(* Logix 5000 project; controller PLC_MCC1300_75F1 vendor 1 type 14 code 166 rev 32.11; software revision 32.04; part 8 of 83 *)

        .rgxMan.4   // Run both
        .rgxMan.5   // Reverse both
        .dErrorCode2   // Error code M2
        .xSensorPresence1   // M403.P115B1.Synchro photocell / start count {x|x|x|x|O}
        .xSensorPresence2   // M403.P115B2.Synchro photocell / start count {x|x|x|x|O}
   M311_HMW : MAC_Conveyor_HMW;
        .dParam_1_cmm   // Positioning offset 1 [mm] {mm/100|mm|-50|+50|M}
        .dParam_2_cmm   // Positioning offset 2 [mm] {mm/100|mm|-50|+50|M}
        .rgxMan.0   // Run M1
        .rgxMan.1   // Reverse M1
        .rgxMan.2   // Run M2
        .rgxMan.3   // Reverse M2
        .rgxMan.4   // Run both
        .rgxMan.5   // Reverse both
   M311_M1_DR : AXIS_CIP_DRIVE; {access Read Only}
   M311_M1_DR_IN_MAJ : MOTION_INSTRUCTION := (FLAGS := 570425344, DN := 1); {access None}
   M311_M1_DR_IN_MAM : MOTION_INSTRUCTION := (FLAGS := 704643072, DN := 1, PC := 1); {access None}
   M311_M1_DR_IN_MAR : MOTION_INSTRUCTION := (FLAGS := 167772160, PC := 1); {access None}
   M311_M1_DR_IN_MAS : MOTION_INSTRUCTION := (FLAGS := -1442840576, EN := 1, DN := 1, PC := 1); {access None}
   M311_M1_DR_IN_MCD : MOTION_INSTRUCTION := (FLAGS := 570425344, DN := 1); {access None}
   M311_M1_DR_IN_MRP : MOTION_INSTRUCTION := (FLAGS := 536870912, DN := 1, STATUS := 2, STATE := 3); {access None}
   M311_M1_DR_MAFR : MOTION_INSTRUCTION := (FLAGS := 301989888, ER := 1, ERR := 11); {access None}
   M311_M1_DR_MDR : MOTION_INSTRUCTION := (FLAGS := -1845493760, EN := 1, ER := 1, ERR := 11); {access None}
   M311_M1_DR_MSF : MOTION_INSTRUCTION := (FLAGS := 570425344, DN := 1, STATUS := 2, STATE := 1); {access None}
   M311_M1_DR_MSO : MOTION_INSTRUCTION := (FLAGS := -1610612736, EN := 1, DN := 1, STATE := 1); {access None}
   M311_M1_DR_OUT_MAJ : MOTION_INSTRUCTION := (FLAGS := 570425344, DN := 1); {access None}
   M311_M1_DR_OUT_MAM : MOTION_INSTRUCTION := (FLAGS := 704643072, DN := 1, PC := 1); {access None}
   M311_M1_DR_OUT_MAR : MOTION_INSTRUCTION := (FLAGS := 671088640, DN := 1, PC := 1, STATE := 1); {access None}
   M311_M1_DR_OUT_MAS : MOTION_INSTRUCTION := (FLAGS := -1442840576, EN := 1, DN := 1, PC := 1); {access None}
   M311_M1_DR_OUT_MCD : MOTION_INSTRUCTION := (FLAGS := 570425344, DN := 1); {access None}
   M311_M1_DR_OUT_MRP : MOTION_INSTRUCTION := (FLAGS := 536870912, DN := 1, STATUS := 2, STATE := 3); {access None}
   M311_SpaceConv_Utilities : SpaceConv_Utilities := (CONST_dSyncMode := 1, CONST_dSyncroPhWindow_cmm := 450000, CONST_dConveyorLength_cmm := 800000, CONST_dConveyorWidth_cmm := 400000, CONST_dPresetFeedbackTime_ms := 500, CONST_rAcceleration_ms2 := 1.2, CONST_rDeceleration_ms2 := 1.2, CONF_MD1_dScan_ms := 20, CONF_MD2_MD3_dPrstPos_cmm := -390000, CONF_MD4_MD6_dLength_cmm := 365800, CONF_MD7_dOffset_cmm := 50000, ST_dStopLoadForseen_cmm := 620000, ST_dRealSpeed_mm_min := 90000, ST_rStepAdvancementH := 3000.0, ST_rStepAdvancementT := 3000.0, O_xPlateSynchronized := 1, O_dCountFeedbackTime_ms := 500, O_dPresetLoadUnload_cmm := -126300);
   M311_SpaceConvUtilities : SpaceConv_Utilities; {access Read Only}
   M311_TON_Synchro_timeout : TIMER; {access Read Only}
   M311_xOS_SentToCullet : BOOL; {access Read Only}
   M311_xPlateCullet : BOOL; {access Read Only}
   M311_xSendCulletReqActive : BOOL; {access Read Only}
   M311_xSensorTimeout : BOOL; {access Read Only}
   M311A : MAC_Rotator := (ST_xCleaningConditionOK := 1, ST_xConditionOKStopCycle := 1, ST_xEnableControlError := 1, INPUT_rRotatorPosition_cdeg := 26999.898, INPUT_xConditionToDescent := 1, INPUT_xLowPosition := 1, INPUT_xLocalSafetySwitchRotation := 1, INPUT_xProtectionMotorLifting := 1, INPUT_xProtectionMotorRotation := 1, tmON_DelayFrameUP.PRE := 100, tmON_DelayRotatorInRun.PRE := 300, tmOF_DriveEnable.PRE := 20000, tmOF_DriveEnable.ACC := 20000, tmON_FeedbackTimeOutLifting.PRE := 1000, tmON_FeedbackTimeOutRotation.PRE := 1000, tmON_FramePosError.PRE := 2500, tmON_RotatePosError.PRE := 10000, tmON_RotatePosError.ACC := 2040, tmON_RotatePosError.EN := 1, tmON_RotatePosError.TT := 1, tmON_PresetEncoder.PRE := 3000, tmON_DelayBrakeON.PRE := 200); {access None}
        .OUTPUT_xDescent   // P253KA4.Descent frame
        .PH_x.0   // Rise frame
        .PH_x.12   // Counterclockwise rotation
        .PH_x.4   // Descent frame
        .PH_x.8   // Clockwise totation
        .OUTPUT_xRise   // P253KA3.Lifting frame
        .INPUT_xLowPosition   // P56KA2.Frame to low position
        .INPUT_xFeedbackLifting   // P56KM1/2.Feedback lifting chassis
        .INPUT_xHighPosition   // P56KA1.Frame to high position
        .INPUT_xProtectionMotorLifting   // P56QM1.Protection lifting frame
   M311A_ALM : MAC_Rotator_ALM;
        .rgxStoppingFault_M[0].0   // Z401.M311A.Protection motor rotation
        .rgxStoppingFault_M[0].1   // Z401.M311A.Drive Error
        .rgxStoppingFault_M[0].11   // Z401.M311A.Frame lifting position error
        .rgxStoppingFault_M[0].2   // Z401.M311A.Drive feedback error
        .rgxStoppingFault_M[0].20   // Z401.M311A.Drive not ready
        .rgxStoppingFault_M[0].3   // Z401.M311A.Rotation position error
        .rgxStoppingFault_M[0].8   // Z401.M311A.Protection lifting frame
        .rgxStoppingFault_M[0].9   // Z401.M311A.Feedback lifting chassis
   M311A_Data : UDT_Convoy_SL;
   M311A_HMR : MAC_Rotator_HMR := (xLowPosition := 1, dState := 1, dActualAngle_cdeg := 27000);
        .rgxMan.0   // Rise
        .rgxMan.1   // Descent
        .rgxMan.10   // Clockwise rotation jog
        .rgxMan.11   // Counter Clockwise rotation jog
        .rgxMan.14   // Enable brake release
        .rgxMan.15   // Disable brake release
        .rgxMan.8   // Clockwise rotation
        .rgxMan.9   // Counter Clockwise rotation
   M311A_HMW : MAC_Rotator_HMW := (xPresetEnc := 1, dLowSpeed_deg_s := 40, dLowRamp_deg_s2 := 50, dHighSpeed_deg_s := 50, dHighRamp_deg_s2 := 60, dJogSpeed_deg_s := 12);
        .rgxMan.0   // Rise
        .rgxMan.1   // Descent
        .rgxMan.10   // Clockwise rotation jog
        .rgxMan.11   // Counterclockwise rotation jog
        .rgxMan.14   // Enable brake release
        .rgxMan.15   // Disable brake release
        .rgxMan.8   // Clockwise rotation
        .rgxMan.9   // Counterclockwise rotation
   M311A_M1_DR : AXIS_CIP_DRIVE; {access Read Only}
   M311A_M1_DR_IN_MAJ : MOTION_INSTRUCTION := (FLAGS := 570425344, DN := 1); {access None}
   M311A_M1_DR_IN_MAM : MOTION_INSTRUCTION := (FLAGS := 704643072, DN := 1, PC := 1); {access None}
   M311A_M1_DR_IN_MAS : MOTION_INSTRUCTION := (FLAGS := -1442840576, EN := 1, DN := 1, PC := 1); {access None}
   M311A_M1_DR_MAFR : MOTION_INSTRUCTION := (FLAGS := 301989888, ER := 1, ERR := 11); {access None}
   M311A_M1_DR_MAH : MOTION_INSTRUCTION := (FLAGS := 671088640, DN := 1, PC := 1, STATE := 17); {access None}
   M311A_M1_DR_MSF : MOTION_INSTRUCTION := (FLAGS := -1610612736, EN := 1, DN := 1, STATUS := 2, STATE := 1); {access None}
   M311A_M1_DR_MSO : MOTION_INSTRUCTION := (FLAGS := 536870912, DN := 1, STATE := 1); {access None}
   M311A_M1_DR_OUT_MAJ : MOTION_INSTRUCTION := (FLAGS := 570425344, DN := 1); {access None}
   M311A_M1_DR_OUT_MAM : MOTION_INSTRUCTION := (FLAGS := 704643072, DN := 1, PC := 1); {access None}
   M311A_M1_DR_OUT_MAS : MOTION_INSTRUCTION := (FLAGS := -1442840576, EN := 1, DN := 1, PC := 1); {access None}
   M311A_MAM_IP_TOFF : TIMER; {access Read Only}
   M311A_rLastPosition : REAL; {access Read Only}
   M311A_TmON1 : TIMER; {access Read Only}
   M311M312_OffsetBaricentre_cmm : DINT; {access Read Only}
   M312 : MAC_Conveyor_Single := (ST_xCleaningConditionOK := 1, ST_xPlatePresence := 1, ST_xConditionOKStopCycle := 1, ST_xOutputEnable := 1, ST_xIdPlatePresence := 1, ST_xWaitStopNextMachine := 1, ST_xEnableControlError := 1, ST_xPlateSynchronized := 1, ST_xSafetyMovement := 1, OSR_xSynchroPhotocellTail := 1, INPUT_xSquaringPhotocell_4 := 1, INPUT_xLowPositionSquaring_1 := 1, INPUT_xHighPositionPopup_1 := 1, INPUT_xHighPositionPopup_2 := 1, INPUT_xDriveReady_M1 := 1, INPUT_xLocalSafetySwitch_M1 := 1, INPUT_xMotorThermalProbe_M1 := 1, INPUT_xProtectionMotor_M1 := 1, INPUT_xDriveReady_M2 := 1, INPUT_xLocalSafetySwitch_M2 := 1, INPUT_xMotorThermalProbe_M2 := 1, INPUT_xProtectionMotor_M2 := 1, INPUT_xDriveFeedback_M3 := 1, INPUT_xDriveReady_M3 := 1, INPUT_xLocalSafetySwitch_M3 := 1, INPUT_xMotorThermalProbe_M3 := 1, INPUT_xProtectionMotor_M3 := 1, INPUT_xDriveReady_M4 := 1, INPUT_xLocalSafetySwitch_M4 := 1, INPUT_xMotorThermalProbe_M4 := 1, INPUT_xProtectionMotor_M4 := 1, INPUT_xProtectionLiftingFrame_1 := 1, INPUT_xProtectionLiftingFrame_2 := 1, INPUT_xFeedbackVentilation_1 := 1, INPUT_xFeedbackVentilation_2 := 1, OUTPUT_xDriveEnable_M1 := 1, OUTPUT_xDriveEnable_M2 := 1, OUTPUT_xDriveEnable_M3 := 1, OUTPUT_xDriveEnable_M4 := 1, OUTPUT_xFunCommand_1 := 1, OUTPUT_xFunCommand_2 := 1, AUX_dPresetStopLoad_cmm := 372333, AUX_dPresetStopUnload_cmm := 441667, AUX_dAccSpace_cmm := 41667, AUX_dDecSpace_cmm := 41667, AUX_dReqSpeed_mm_min := 60000, AUX_dAbsPosTarget_M3_cmm := 195500, AUX_dAbsPosTarget_M4_cmm := 195500, AUX_dQtaLites := 1, tmON_FeedbackTimeOut_M1.PRE := 2000, tmOF_DriveEnable_M1.PRE := 30000, tmOF_DriveEnable_M1.ACC := 540, tmOF_DriveEnable_M1.TT := 1, tmOF_DriveEnable_M1.DN := 1, tmOF_PowerSaving_M1.EN := 1, tmOF_PowerSaving_M1.DN := 1, tmON_FeedbackTimeOut_M2.PRE := 2000, tmOF_DriveEnable_M2.PRE := 30000, tmOF_DriveEnable_M2.ACC := 540, tmOF_DriveEnable_M2.TT := 1,
        tmOF_DriveEnable_M2.DN := 1, tmON_FeedbackTimeOut_M3.PRE := 2000, tmOF_DriveEnable_M3.PRE := 30000, tmOF_DriveEnable_M3.ACC := 540, tmOF_DriveEnable_M3.TT := 1, tmOF_DriveEnable_M3.DN := 1, tmON_FeedbackTimeOut_M4.PRE := 2000, tmOF_DriveEnable_M4.PRE := 30000, tmOF_DriveEnable_M4.ACC := 540, tmOF_DriveEnable_M4.TT := 1, tmOF_DriveEnable_M4.DN := 1, tmON_AuxFunction1.PRE := 5000, tmON_AuxFunction1.EN := 1, tmON_AuxFunction1.DN := 1, tmON_AuxFunction2.PRE := 2200, tmON_AuxFunction3.PRE := 2200, tmON_AuxFunction4.PRE := 15000, tmON_AuxFunction5.PRE := 3000, tmON_AuxFunction6.PRE := 15000, tmON_AuxFunction7.PRE := 3600000, tmON_AuxFunction8.PRE := 40000, tmON_AuxFunction9.PRE := 20000, TmON[0].PRE := 3000, TmON[1].PRE := 1000, TmON[1].ACC := 1019, TmON[2].PRE := 5000, TmON[6].PRE := 5000, TmON[6].EN := 1, TmON[6].DN := 1, TmON[11].PRE := 2000, TmON[12].PRE := 2000, TmON[13].PRE := 2000, TmON[14].PRE := 2000, tmOF_MCD_M1.ACC := 20, tmOF_MCD_M2.ACC := 20, tmOF_MCD_M3.ACC := 20, tmOF_MCD_M4.ACC := 20); {access None}
        .INPUT_xSquaringPhotocell_1   // P406B1.Squaring frontal photocell - Right
        .INPUT_xMotorThermalProbe_M2   // M2.P404BT2.Motor thermal probe
        .INPUT_xLowPositionPopup_1   // P63KA2.M5.Low position popup
        .INPUT_xLowPositionSquaring_1   // P405SQ2.Low position squaring
        .INPUT_xMotorThermalProbe_M1   // M1.P404BT1.Motor thermal probe
        .INPUT_xHighPositionPopup_1   // P63KA1.M5.High position popup
        .INPUT_xSquaringPhotocell_2   // P406B2.Squaring frontal photocell - Left
        .INPUT_xHighPositionPopup_2   // P64KA1.M6.High position popup
        .PH_x.0   // Load (from M311)
        .PH_x.10   // Load (from M409)
        .PH_x.11   // End load (from M409)
        .PH_x.12   // Unload (to M311)
        .PH_x.13   // End unload (to M311)
        .PH_x.15   // End unload (to M409)
        .PH_x.16   // Rise popup
        .PH_x.19   // End rise popup
        .PH_x.20   // Descent popup
        .PH_x.23   // End descent popup
        .PH_x.24   // Reset counter position
        .PH_x.26   // Lateral positioning (M3-M4)
        .PH_x.27   // End lateral positioning (M3-M4)
        .PH_x.28   // Lateral squaring
        .PH_x.29   // End lateral squaring
        .PH_x.30   // Lateral traction recovery (M3-M4)
        .PH_x.31   // End lateral traction recovery (M3-M4)
        .PH_x.4   // Frontal squaring (run fwd + rise squaring)
        .PH_x.5   // End frontal sqauring
        .PH_x.7   // End load (from M311)
        .PH_x.8   // Unload (to M409)
        .INPUT_xMotorThermalProbe_M3   // M3.P405BT3.Motor thermal probe
        .INPUT_xLowPositionPopup_2   // P64KA2.M6.Low position popup
        .INPUT_xSquaringPhotocell_3   // P405B1.Squaring lateral photocell - Right
        .INPUT_xHighPositionSquaring_1   // P405SQ1.High position squaring
        .INPUT_xSquaringPhotocell_4   // P405B2.Squaring lateral photocell - Left
        .INPUT_xHighPositionSquaring_2   // P405SQ11.High position squaring
        .ST_xAux1   // Ready to unload on backward conveyor
        .INPUT_xLowPositionSquaring_2   // P405SQ12.Low position squaring
   M312_ALM : MAC_Conveyor_ALM;
        .rgdFaultCode_M[0]   // Drive fault code M1
        .rgdFaultCode_M[1]   // Drive fault code M2
        .rgxStoppingFault[0].0   // Z401.M312-M1.Positioning error
        .rgxStoppingFault[0].1   // Z401.M312-M1.Plate not synchronized
        .rgxStoppingFault[0].10   // Z401.M312-M2.Error position frontal squaring
        .rgxStoppingFault[0].11   // Z401.M312-M2.Timeout frontal squaring
        .rgxStoppingFault[0].12   // Z401.M312-M2.Lugs position sensors fault
        .rgxStoppingFault[0].13   // Z401.M312.Timeout movement popup 1
        .rgxStoppingFault[0].14   // Z401.M312.Timeout movement popup 1
        .rgxStoppingFault[0].16   // Z401.M312-M3.Positioning error
        .rgxStoppingFault[0].18   // Z401.M312-M3.Error position popup
        .rgxStoppingFault[0].19   // Z401.M312-M3.Error position lateral squaring
        .rgxStoppingFault[0].2   // Z401.M312-M1.Error position frontal squaring
        .rgxStoppingFault[0].20   // Z401.M312-M3.Timeout lateral squaring
        .rgxStoppingFault[0].21   // Z401.M312.Protection lifting popup 1
        .rgxStoppingFault[0].22   // Z401.M312.Protection lifting popup 2
        .rgxWarning[0].10   // Z401.M312_M2.Plate not synchronized
        .rgxStoppingFault[0].3   // Z401.M312-M1.Timeout frontal squaring
        .rgxStoppingFault[0].4   // Z401.M312-M1.Lugs position sensors fault
        .rgxStoppingFault[0].5   // Z401.M312.Popup 1 position error
        .rgxStoppingFault[0].6   // Z401.M312.Popup 2 position error
        .rgxStoppingFault[0].8   // Z401.M312-M2.Positioning error
        .rgxStoppingFault[0].9   // Z401.M312-M2.Plate not synchronized
        .rgxStoppingFault_M[0].0   // Z401.M312-M1.Protection motor rotation
        .rgxStoppingFault_M[0].1   // Z401.M312-M1.Drive error
        .rgxStoppingFault_M[0].10   // Z401.M312-M2.Drive feedback error
        .rgxStoppingFault_M[0].11   // Z401.M312-M2.Local safety switch
        .rgxStoppingFault_M[0].12   // Z401.M312-M2.Motor thermal probe
        .rgxStoppingFault_M[0].13   // Z401.M312-M2.Braking resistor anomaly
        .rgxStoppingFault_M[0].14   // Z401.M312-M2.Drive not ready
        .rgxStoppingFault_M[0].16   // Z401.M312-M3.Protection motor rotation
        .rgxStoppingFault_M[0].17   // Z401.M312-M3.Drive error
        .rgxStoppingFault_M[0].18   // Z401.M312-M3.Drive feedback error
        .rgxStoppingFault_M[0].19   // Z401.M312-M3.Local safety switch
        .rgxStoppingFault_M[0].2   // Z401.M312-M1.Drive feedback error
        .rgxStoppingFault_M[0].20   // Z401.M312-M3.Motor thermal probe
        .rgxStoppingFault_M[0].21   // Z401.M312-M3.Drive not ready
        .rgxStoppingFault_M[0].3   // Z401.M312-M1.Local safety switch
        .rgxStoppingFault_M[0].4   // Z401.M312-M1.Motor thermal probe
        .rgxStoppingFault_M[0].5   // Z401.M312-M1.Braking resistor anomaly
        .rgxStoppingFault_M[0].6   // Z401.M312-M1.Drive not ready
        .rgxStoppingFault_M[0].8   // Z401.M312-M2.Protection motor rotation
        .rgxStoppingFault_M[0].9   // Z401.M312-M2.Drive error
        .rgxWarning[0].0   // Z401.M312_M1.Plate not synchronized
        .rgxWarning[0].1   // Z401.M312_M1.Positioning error
        .rgxWarning[0].11   // Z401.M312_M2.Positioning error
        .rgxWarning[0].21   // Z401.M312_M3.Lateal positioning error
        .rgxWarning[0].25   // Z401.M312.Timeout frontal squaring
        .rgxWarning[0].26   // Z401.M312.Timeout lateral squaring
   M312_AlmTimer1 : TIMER; {access Read Only}
   M312_AlmTimer2 : TIMER; {access Read Only}
   M312_Data : UDT_Convoy_SL;
        .rgtCap[0].rgxRequest.0   // Frontal squaring request
        .rgtCap[0].rgxRequest.1   // Lateral squaring request
        .rgtCap[0].rgxRequest.2   // Y adjust position request
        .rgtCap[0].rgxRequest.3   // Y measure request
        .rgtCap[0].rgxDone.0   // Frontal squaring done
        .rgtCap[0].rgxDone.1   // Lateral squaring done
        .rgtCap[0].rgxDone.2   // Y adjust position done
        .rgtCap[0].rgxDone.3   // Y measure done
   M312_dSlowingSquaringQuote : DINT; {access Read Only}
   M312_dTractionRecovery_M3 : DINT; {access Read Only}
   M312_dTractionRecovery_M4 : DINT; {access Read Only}
   M312_HMR : MAC_Conveyor_HMR := (xSensorPresence4 := 1, xHighPositionPopup1 := 1, xHighPositionPopup2 := 1, xLowPositionSquaring1 := 1, xLowPositionSquaring2 := 1, xIdPlatePresence := 1, dState1 := 1, dState2 := 1, dState3 := 1, dState4 := 1, dStateSensor1 := 1, dStateSensor2 := 1, dStateSensor3 := 1, dStateSensor4 := 1, dStateSensor5 := 1, dStateSensor6 := 1);
        .xSensorPresence5   // P115/3.Start count photocell {x|x|x|x|O}
        .xHighPositionPopup2   // P64KA1.M6.High position popup {x|x|x|x|O}
        .dErrorCode1   // Error code M1
        .xHighPositionPopup1   // P63KA1.M5.High position popup {x|x|x|x|O}
        .rgxMan.0   // Run M1
        .rgxMan.1   // Reverse M1
        .rgxMan.10   // Rise popup 1
        .rgxMan.11   // Descent popup 1
        .rgxMan.12   // Rise popup 2
        .rgxMan.13   // Descent popup 2
        .rgxMan.14   // Rise all popups
        .rgxMan.15   // Descent all popups
        .rgxMan.16   // Rise frontal squaring 1
        .rgxMan.17   // Descent frontal squaring 1
        .rgxMan.18   // Rise frontal squaring 2
        .rgxMan.19   // Descent frontal squaring 2
        .rgxMan.2   // Run M2
        .rgxMan.20   // Rise all frontal squaring
        .rgxMan.21   // Descent all frontal squaring
        .rgxMan.3   // Reverse M2
        .rgxMan.4   // Run M3
        .rgxMan.5   // Reverse M3
        .rgxMan.6   // Run M4
        .rgxMan.7   // Reverse M4
        .dState3   // State M3 (1=No anomaly; 3=Run; 4=Reverse; 7=Anomaly)
        .xHighPositionSquaring1   // P405SQ1.High position frontal squaring M1 {x|x|x|x|O}
        .dErrorCode2   // Error code M2
        .xSensorPresence6   // P115/4.Start count photocell {x|x|x|x|O}
        .xSensorPresence4   // P404B1.SlowDown photocell frontal squaring left {x|x|x|x|O}
        .xLowPositionPopup1   // P63KA2.M5.Low position popup {x|x|x|x|O}
        .xHighPositionSquaring2   // P405SQ11.High position frontal squaring M2 {x|x|x|x|O}
        .dState2   // State M2 (1=No anomaly; 3=Run; 4=Reverse; 7=Anomaly)
        .dErrorCode4   // Error code M4
        .xSensorPresence3   // P404B1.SlowDown photocell frontal squaring right {x|x|x|x|O}
        .dState1   // State M1 (1=No anomaly; 3=Run; 4=Reverse; 7=Anomaly)
        .dState4   // State M4 (1=No anomaly; 3=Run; 4=Reverse; 7=Anomaly)
        .xLowPositionSquaring2   // P405SQ12.Low position frontal squaring M2 {x|x|x|x|O}
        .xLowPositionSquaring1   // P405SQ2.Low position frontal squaring M1 {x|x|x|x|O}
        .xLowPositionPopup2   // P64KA2.M6.Low position popup {x|x|x|x|O}
        .xSensorPresence1   // P405B1.SlowDown photocell lateral squaring right {x|x|x|x|O}
        .dErrorCode3   // Error code M3
        .xSensorPresence2   // P405B2.SlowDown photocell lateral squaring left {x|x|x|x|O}
   M312_HMW : MAC_Conveyor_HMW := (dParam_3_cmm := 4000, dParam_5_ms := 3000, dParam_6_ms := 4000, dParam_7_ms := 2200, dParam_8_ms := 5000);
        .dParam_4_cmm   // Lateral squaring space {mm/100|mm|0|500|M}
        .dParam_1_cmm   // Positioning offset 1 {mm/100|mm|-50|+50|M}
        .dParam_3_cmm   // Frontal squaring space {mm/100|mm|0|500|M}
        .dParam_6_ms   // Squaring frontal time 2 {ms|s|0|5|M}
        .dParam_2_cmm   // Positioning offset 2 {mm/100|mm|-50|+50|M}
        .dParam_8_ms   // Squaring lateral time 2 {ms|s|0|5|M}
        .rgxMan.0   // Run M1
        .rgxMan.1   // Reverse M1
        .rgxMan.10   // Rise popup 2
        .rgxMan.11   // Descent popup 2
        .rgxMan.12   // Rise all popups
        .rgxMan.13   // Descent all popups
        .rgxMan.14   // Run both (M1-2)
        .rgxMan.15   // Reverse both (M1-2)
        .rgxMan.16   // Rise frontal squaring 1
        .rgxMan.17   // Descent frontal squaring 1
        .rgxMan.18   // Rise frontal squaring 2
        .rgxMan.19   // Descent frontal squaring 2
        .rgxMan.2   // Run M2
        .rgxMan.20   // Rise all frontal squaring
        .rgxMan.21   // Descent all frontal squaring
        .rgxMan.3   // Reverse M2
        .rgxMan.4   // Run M3
        .rgxMan.5   // Reverse M3
        .rgxMan.6   // Run M4
        .rgxMan.7   // Reverse M4
        .rgxMan.8   // Rise popup 1
        .rgxMan.9   // Descent popup 1
        .dParam_7_ms   // Squaring lateral time 1 {ms|s|0|5|M}
        .dParam_5_ms   // Squaring frontal time 1 {ms|s|0|5|M}
   M312_M1_DR_IN_MAJ : MOTION_INSTRUCTION := (FLAGS := 570425344, DN := 1); {access None}
   M312_M1_DR_IN_MAM : MOTION_INSTRUCTION := (FLAGS := 33554432); {access None}
   M312_M1_DR_IN_MAR : MOTION_INSTRUCTION := (FLAGS := 33554432); {access None}
   M312_M1_DR_IN_MAS : MOTION_INSTRUCTION := (FLAGS := -1442840576, EN := 1, DN := 1, PC := 1); {access None}
   M312_M1_DR_IN_MCD : MOTION_INSTRUCTION := (FLAGS := 570425344, DN := 1); {access None}
   M312_M1_DR_IN_MRP : MOTION_INSTRUCTION := (FLAGS := 33554432); {access None}
   M312_M1_DR_MAFR : MOTION_INSTRUCTION := (FLAGS := 301989888, ER := 1, ERR := 11); {access None}
   M312_M1_DR_MDR : MOTION_INSTRUCTION := (FLAGS := -1845493760, EN := 1, ER := 1, ERR := 11); {access None}
   M312_M1_DR_MSF : MOTION_INSTRUCTION := (FLAGS := 570425344, DN := 1, STATUS := 2, STATE := 1); {access None}
   M312_M1_DR_MSO : MOTION_INSTRUCTION := (FLAGS := -1610612736, EN := 1, DN := 1, STATE := 1); {access None}
   M312_M1_DR_OUT_MAJ : MOTION_INSTRUCTION := (FLAGS := 570425344, DN := 1); {access None}
   M312_M1_DR_OUT_MAM : MOTION_INSTRUCTION := (FLAGS := 33554432); {access None}
   M312_M1_DR_OUT_MAR : MOTION_INSTRUCTION := (FLAGS := 33554432); {access None}
   M312_M1_DR_OUT_MAS : MOTION_INSTRUCTION := (FLAGS := -1442840576, EN := 1, DN := 1, PC := 1); {access None}
   M312_M1_DR_OUT_MCD : MOTION_INSTRUCTION := (FLAGS := 570425344, DN := 1); {access None}
   M312_M1_DR_OUT_MRP : MOTION_INSTRUCTION := (FLAGS := 33554432); {access None}
   M312_M1_DR_R1 : AXIS_CIP_DRIVE; {access Read Only}
   M312_M2_AUX_ReqSpeed_mm_min : DINT; {access Read Only}
   M312_M2_ChangeSpeed : BOOL; {access Read Only}
   M312_M2_DR_IN_MAJ : MOTION_INSTRUCTION := (FLAGS := 570425344, DN := 1); {access None}
   M312_M2_DR_IN_MAM : MOTION_INSTRUCTION := (FLAGS := 33554432); {access None}
   M312_M2_DR_IN_MAR : MOTION_INSTRUCTION := (FLAGS := 33554432); {access None}
   M312_M2_DR_IN_MAS : MOTION_INSTRUCTION := (FLAGS := 704643072, DN := 1, PC := 1); {access None}
   M312_M2_DR_IN_MCD : MOTION_INSTRUCTION := (FLAGS := 301989888, ER := 1, ERR := 23); {access None}
   M312_M2_DR_IN_MRP : MOTION_INSTRUCTION := (FLAGS := 536870912, DN := 1, STATUS := 2, STATE := 3); {access None}
   M312_M2_DR_MAFR : MOTION_INSTRUCTION := (FLAGS := 301989888, ER := 1, ERR := 11); {access None}
   M312_M2_DR_MDR : MOTION_INSTRUCTION := (FLAGS := -1845493760, EN := 1, ER := 1, ERR := 11); {access None}
   M312_M2_DR_MSF : MOTION_INSTRUCTION := (FLAGS := 570425344, DN := 1, STATUS := 2, STATE := 1); {access None}
   M312_M2_DR_MSO : MOTION_INSTRUCTION := (FLAGS := -1610612736, EN := 1, DN := 1, STATE := 1); {access None}
   M312_M2_DR_OUT_MAJ : MOTION_INSTRUCTION := (FLAGS := 570425344, DN := 1); {access None}
   M312_M2_DR_OUT_MAM : MOTION_INSTRUCTION := (FLAGS := 33554432); {access None}
   M312_M2_DR_OUT_MAR : MOTION_INSTRUCTION := (FLAGS := 33554432); {access None}
   M312_M2_DR_OUT_MAS : MOTION_INSTRUCTION := (FLAGS := 704643072, DN := 1, PC := 1); {access None}
   M312_M2_DR_OUT_MCD : MOTION_INSTRUCTION := (FLAGS := 301989888, ER := 1, ERR := 23); {access None}
   M312_M2_DR_OUT_MRP : MOTION_INSTRUCTION := (FLAGS := 536870912, DN := 1, STATUS := 2, STATE := 3); {access None}
   M312_M2_DR_R2 : AXIS_CIP_DRIVE; {access Read Only}
   M312_M2_ReqSpeed_mm_min : DINT; {access Read Only}
   M312_M3_AUX_ReqSpeed_mm_min : DINT; {access Read Only}
   M312_M3_ChangeSpeed : BOOL; {access Read Only}
   M312_M3_DR_IN_MAJ : MOTION_INSTRUCTION := (FLAGS := 570425344, DN := 1); {access None}
   M312_M3_DR_IN_MAM : MOTION_INSTRUCTION := (FLAGS := -1509949440, EN := 1, DN := 1, IP := 1); {access None}
   M312_M3_DR_IN_MAR : MOTION_INSTRUCTION := (FLAGS := 33554432); {access None}
   M312_M3_DR_IN_MAS : MOTION_INSTRUCTION := (FLAGS := 704643072, DN := 1, PC := 1); {access None}
   M312_M3_DR_IN_MCD : MOTION_INSTRUCTION := (FLAGS := 570425344, DN := 1); {access None}
   M312_M3_DR_IN_MRP : MOTION_INSTRUCTION := (FLAGS := 536870912, DN := 1, STATUS := 2, STATE := 3); {access None}
   M312_M3_DR_L : AXIS_CIP_DRIVE; {access Read Only}
   M312_M3_DR_MAFR : MOTION_INSTRUCTION := (FLAGS := 301989888, ER := 1, ERR := 11); {access None}
   M312_M3_DR_MDR : MOTION_INSTRUCTION := (FLAGS := -1845493760, EN := 1, ER := 1, ERR := 11); {access None}
   M312_M3_DR_MSF : MOTION_INSTRUCTION := (FLAGS := 570425344, DN := 1, STATUS := 2, STATE := 1); {access None}
   M312_M3_DR_MSO : MOTION_INSTRUCTION := (FLAGS := -1610612736, EN := 1, DN := 1, STATE := 1); {access None}
   M312_M3_DR_OUT_MAJ : MOTION_INSTRUCTION := (FLAGS := 570425344, DN := 1); {access None}
   M312_M3_DR_OUT_MAM : MOTION_INSTRUCTION := (FLAGS := -1509949440, EN := 1, DN := 1, IP := 1);
   M312_M3_DR_OUT_MAR : MOTION_INSTRUCTION := (FLAGS := 33554432); {access None}
   M312_M3_DR_OUT_MAS : MOTION_INSTRUCTION := (FLAGS := 704643072, DN := 1, PC := 1); {access None}
   M312_M3_DR_OUT_MCD : MOTION_INSTRUCTION := (FLAGS := 570425344, DN := 1); {access None}
   M312_M3_DR_OUT_MRP : MOTION_INSTRUCTION := (FLAGS := 536870912, DN := 1, STATUS := 2, STATE := 3); {access None}
   M312_M3_ReqSpeed_mm_min : DINT; {access Read Only}
   M312_M3_xOSR_LatSquarFtc : BOOL; {access Read Only}
   M312_SpaceConv_Utilities : SpaceConv_Utilities := (CONST_dSyncMode := 1, CONST_dSyncroPhWindow_cmm := 450000, CONST_dConveyorLength_cmm := 800000, CONST_dConveyorWidth_cmm := 400000, CONST_dPresetFeedbackTime_ms := 500, CONST_rAcceleration_ms2 := 1.2, CONST_rDeceleration_ms2 := 1.2, CONF_MD1_dScan_ms := 20, CONF_MD2_MD3_dPrstPos_cmm := -390000, CONF_MD4_MD6_dLength_cmm := 365800, CONF_MD7_dOffset_cmm := 50000, ST_dStopLoadForseen_cmm := 620000, ST_dRealSpeed_mm_min := 90000, ST_rStepAdvancementH := 3000.0, ST_rStepAdvancementT := 3000.0, O_xPlateSynchronized := 1, O_dCountFeedbackTime_ms := 500, O_dPresetLoadUnload_cmm := -126300);
   M312_TimerAlm3 : TIMER; {access Read Only}
   M312_TON_FrontSquarLeft_timeout : TIMER; {access Read Only}
   M312_TON_FrontSquarRight_timeout : TIMER; {access Read Only}
   M312_TON_LatSquarLeft_timeout : TIMER; {access Read Only}
   M312_TON_LatSquarRight_timeout : TIMER; {access Read Only}
   M312_TON_Load : TIMER; {access Read Only}
   M312_TON_Synchro_timeout : TIMER; {access Read Only}
   M312_xEnableTractionRecovering : BOOL; {access Read Only}
   M312_xFrontLeftTimeout : BOOL; {access Read Only}
   M312_xFrontRightTimeout : BOOL; {access Read Only}
   M312_xLateralTractionRecovered : BOOL; {access Read Only}
   M312_xLatLeftTimeout : BOOL; {access Read Only}
   M312_xLatRightTimeout : BOOL; {access Read Only}
   M312_xOS_PosReq : BOOL;
   M312_xPlateCullet : BOOL; {access Read Only}
   M312_xSendCulletReqActive : BOOL; {access Read Only}
   M312_xSensorTimeout : BOOL; {access Read Only}
   M315_M1_DR_R1 : AXIS_CIP_DRIVE; {access Read Only}
   M315_M2_DR_R2 : AXIS_CIP_DRIVE; {access Read Only}
   M315_M3_DR_R3 : AXIS_CIP_DRIVE; {access Read Only}
   M315_M4_DR_B1 : AXIS_CIP_DRIVE; {access Read Only}
   M315_M5_DR_B2 : AXIS_CIP_DRIVE; {access Read Only}
   M315_M6_DR_L1 : AXIS_CIP_DRIVE; {access Read Only}
   M315_M7_DR_L2 : AXIS_CIP_DRIVE; {access Read Only}
   M315_xReqStopPrevConvForPos : BOOL; {access Read Only}
   M315A : MAC_Conveyor;
        .PH_x.1   // Load Upstream
        .PH_x.0   // Load
        .PH_x.7   // End load
        .PH_x.8   // Unload
        .PH_x.15   // End unload
        .INPUT_xMotorThermalProbe_M1   // M315A.M1.Q403BT3. Motor thermal probe
        .PH_x.2   // Load Downstream
        .PH_x.5   // End load Upstream
        .PH_x.6   // End load Downstream
        .PH_x.9   // Unload Upstream
        .PH_x.10   // Unload Downstream
        .PH_x.13   // End unload Upstream
        .PH_x.14   // End unload Downstream
        .PH_x.16   // Unpack convoy
        .PH_x.17   // End unpack convoy
        .PH_x.18   // Unpack convoy Upstream
        .PH_x.19   // End unpack convoy Upstream
        .PH_x.21   // End unpack convoy Downstream
        .PH_x.20   // Unpack convoy Downstream
        .PH_x.22   // Stop for unload on main line
        .PH_x.23   // End stop for unload on main line
        .PH_x.28   // Load reentry
        .PH_x.29   // End load reentry
        .PH_x.24   // Stop for unload on main line Upstream
        .PH_x.25   // End stop for unload on main line Upstream
        .PH_x.26   // Stop for unload on main line Downstream
        .PH_x.27   // End stop for unload on main line Downstream
   M315A_ALM : MAC_Conveyor_ALM;
        .rgdFaultCode_M[0]   // Drive fault code
        .rgxStoppingFault_M[0].5   // Z402.M315A-M1.Braking resistor anomaly
        .rgxStoppingFault_M[0].1   // Z402.M315A-M1.Drive error
        .rgxStoppingFault_M[0].6   // Z402.M315A-M1.Drive not ready
        .rgxStoppingFault_M[0].4   // Z402.M315A.M1. Motor thermal probe
        .rgxStoppingFault_M[0].3   // Z402.M315A-M1.Local safety switch
        .rgxStoppingFault_M[0].0   // Z402.M315A-M1.Protection motor rotation
        .rgxStoppingFault_M[0].2   // Z402.M315A-M1.Drive feedback error
        .rgxWarning[0].1   // Z402.M315A.Positioning error
        .rgxWarning[0].0   // Z402.M315A.Q115B1.Plate not synchronized
   M315A_Data : UDT_Convoy_SL;
   M315A_dLastSyncID : DINT; {access Read Only}
   M315A_HMR : MAC_Conveyor_HMR := (xManualCommandEnabled := 1, dState4 := 1);
        .dErrorCode1   // Error code M1
        .rgxMan.0   // Run M1
        .rgxMan.1   // Reverse M1
        .rgxMan.2   // Run M2
        .rgxMan.3   // Reverse M2
        .rgxMan.4   // Run M3
        .rgxMan.5   // Reverse M3
        .dErrorCode2   // Error code M2 (NU)
        .xSensorPresence1   // M501.Q115B1. Sincro phoyocell / start count {x|x|x|xO}
        .dErrorCode3   // Error code M3 (NU)
   M315A_HMW : MAC_Conveyor_HMW;
        .rgxMan.0   // Run M1
        .rgxMan.1   // Reverse M1
        .rgxMan.2   // Run M2
        .rgxMan.3   // Reverse M2
        .rgxMan.4   // Run M3
        .rgxMan.5   // Reverse M3
   M315A_INPUT_xSyncroPhotocell : BOOL; {access Read Only}
   M315A_M1_DR : AXIS_CIP_DRIVE; {access Read Only}
   M315A_M1_DR_IN_MAJ : MOTION_INSTRUCTION := (FLAGS := 570425344, DN := 1); {access None}
   M315A_M1_DR_IN_MAM : MOTION_INSTRUCTION := (FLAGS := 33554432); {access None}
   M315A_M1_DR_IN_MAR : MOTION_INSTRUCTION := (FLAGS := 33554432); {access None}
   M315A_M1_DR_IN_MAS : MOTION_INSTRUCTION := (FLAGS := -1442840576, EN := 1, DN := 1, PC := 1); {access None}
   M315A_M1_DR_IN_MCD : MOTION_INSTRUCTION := (FLAGS := 570425344, DN := 1); {access None}
   M315A_M1_DR_IN_MRP : MOTION_INSTRUCTION := (FLAGS := 33554432); {access None}
   M315A_M1_DR_MAFR : MOTION_INSTRUCTION := (FLAGS := 301989888, ER := 1, ERR := 11); {access None}
   M315A_M1_DR_MDR : MOTION_INSTRUCTION := (FLAGS := -1845493760, EN := 1, ER := 1, ERR := 11); {access None}
   M315A_M1_DR_MSF : MOTION_INSTRUCTION := (FLAGS := 536870912, DN := 1, STATUS := 2, STATE := 1); {access None}
   M315A_M1_DR_MSO : MOTION_INSTRUCTION := (FLAGS := -1577058304, EN := 1, DN := 1, STATE := 1); {access None}
   M315A_M1_DR_OUT_MAJ : MOTION_INSTRUCTION := (FLAGS := 570425344, DN := 1); {access None}
   M315A_M1_DR_OUT_MAM : MOTION_INSTRUCTION := (FLAGS := 33554432); {access None}
   M315A_M1_DR_OUT_MAR : MOTION_INSTRUCTION := (FLAGS := 33554432); {access None}
   M315A_M1_DR_OUT_MAS : MOTION_INSTRUCTION := (FLAGS := -1442840576, EN := 1, DN := 1, PC := 1); {access None}
   M315A_M1_DR_OUT_MCD : MOTION_INSTRUCTION := (FLAGS := 570425344, DN := 1); {access None}
   M315A_M1_DR_OUT_MRP : MOTION_INSTRUCTION := (FLAGS := 33554432); {access None}
   M315A_OSR_xSyncOnLoad : BOOL; {access Read Only}
   M315A_SpaceConv_Utilities : SpaceConv_Utilities := (CONST_dSyncMode := 1, CONST_dSyncroPhWindow_cmm := 450000, CONST_dConveyorLength_cmm := 800000, CONST_dConveyorWidth_cmm := 400000, CONST_dPresetFeedbackTime_ms := 500, CONST_rAcceleration_ms2 := 1.2, CONST_rDeceleration_ms2 := 1.2, CONF_MD1_dScan_ms := 20, CONF_MD2_MD3_dPrstPos_cmm := -390000, CONF_MD4_MD6_dLength_cmm := 365800, CONF_MD7_dOffset_cmm := 50000, ST_dStopLoadForseen_cmm := 620000, ST_dRealSpeed_mm_min := 90000, ST_rStepAdvancementH := 3000.0, ST_rStepAdvancementT := 3000.0, O_xPlateSynchronized := 1, O_dCountFeedbackTime_ms := 500, O_dPresetLoadUnload_cmm := -126300);
   M315A_SpaceConvUtilities : SpaceConv_Utilities; {access Read Only}
   M315A_xSyncOnLoadDone : BOOL; {access Read Only}
   M315B : MAC_Conveyor := (ST_xCleaningConditionOK := 1, ST_xConditionOKStopCycle := 1, ST_xEnableControlError := 1, ST_xSafetyMovement := 1, ST_xAux4 := 1, OSR_xSynchroPhotocellTail := 1, INPUT_xLowPositionPopup_1 := 1, INPUT_xLowPositionPopup_2 := 1, INPUT_xDriveReady_M2 := 1, INPUT_xDriveReady_M3 := 1, INPUT_xLocalSafetySwitch_M3 := 1, INPUT_xProtectionMotor_M3 := 1, INPUT_xDriveReady_M4 := 1, INPUT_xLocalSafetySwitch_M4 := 1, INPUT_xProtectionMotor_M4 := 1, OUTPUT_xDriveEnable_M3 := 1, OUTPUT_xDriveEnable_M4 := 1, AUX_dPresetStopLoad_cmm := 455000, AUX_dPresetStopUnload_cmm := 575000, AUX_dAccSpace_cmm := 41667, AUX_dDecSpace_cmm := 41667, AUX_dReqSpeed_mm_min := 60000, AUX_dPhPosTarget_cmm := 180000, TmON_AxleReadyToMoveDelayed.PRE := 500, tmON_FeedbackTimeOut_M1.PRE := 1500, tmOF_DriveEnable_M1.PRE := 20000, tmOF_DriveEnable_M1.ACC := 6500, tmOF_DriveEnable_M1.TT := 1, tmOF_DriveEnable_M1.DN := 1, tmOF_PowerSaving_M1.PRE := 20000, tmOF_PowerSaving_M1.ACC := 20000, tmOF_PowerSaving_M1.EN := 1, tmOF_PowerSaving_M1.DN := 1, tmON_FeedbackTimeOut_M2.PRE := 1500, tmOF_DriveEnable_M2.PRE := 20000, tmOF_DriveEnable_M2.ACC := 3500, tmOF_PowerSaving_M2.PRE := 20000, tmON_FeedbackTimeOut_M3.PRE := 1500, tmOF_DriveEnable_M3.PRE := 20000, tmOF_DriveEnable_M3.ACC := 6500, tmOF_DriveEnable_M3.TT := 1, tmOF_DriveEnable_M3.DN := 1, tmOF_PowerSaving_M3.PRE := 20000, tmOF_PowerSaving_M3.ACC := 20000, tmON_FeedbackTimeOut_M4.PRE := 1500, tmOF_DriveEnable_M4.PRE := 20000, tmOF_DriveEnable_M4.ACC := 3500, tmOF_DriveEnable_M4.TT := 1, tmOF_DriveEnable_M4.DN := 1, tmOF_MCD_M1.PRE := 200, tmOF_MCD_M1.ACC := 200, tmOF_MCD_M2.PRE := 200, tmOF_MCD_M2.ACC := 200, tmOF_MCD_M3.PRE := 200, tmOF_MCD_M3.ACC := 200, tmOF_MCD_M4.PRE := 200, tmOF_MCD_M4.ACC := 200); {access None}
        .INPUT_xMotorThermalProbe_M2   // M325.M4.P403BT2.Motor thermal probe
        .INPUT_xMotorThermalProbe_M1   // M325.M3.P403BT1.Motor thermal probe
        .PH_x.0   // Load
        .PH_x.1   // Load Upstream
        .PH_x.10   // Unload Downstream
        .PH_x.13   // End unload Upstream
        .PH_x.14   // End unload Downstream
        .PH_x.15   // End unload
        .PH_x.16   // Unpack convoy
        .PH_x.17   // End unpack convoy
        .PH_x.18   // Unpack convoy Upstream
        .PH_x.19   // End unpack convoy Upstream
        .PH_x.2   // Load Downstream
        .PH_x.20   // Unpack convoy Downstream
        .PH_x.21   // End unpack convoy Downstream
        .PH_x.22   // Stop for unload on main line
        .PH_x.23   // End stop for unload on main line
        .PH_x.24   // Stop for unload on main line Upstream
        .PH_x.25   // End stop for unload on main line Upstream
        .PH_x.26   // Stop for unload on main line Downstream
        .PH_x.27   // End stop for unload on main line Downstream
        .PH_x.28   // Load reentry
        .PH_x.29   // End load reentry
        .PH_x.5   // End load Upstream
        .PH_x.6   // End load Downstream
        .PH_x.7   // End load
        .PH_x.8   // Unload
        .PH_x.9   // Unload Upstream
   M315B_ALM : MAC_Conveyor_ALM;
        .rgxStoppingFault_M[0].1   // Z402.M315B-M1.P51AZ1.Drive error
        .rgxStoppingFault_M[0].13   // Z402.M315B-M2.P51AZ1.Local safety switch
        .rgxStoppingFault_M[0].11   // Z402.M315B-M2.P51AZ1.Drive error
        .rgxStoppingFault_M[0].0   // Z402.M315B-M1.P51AZ1.Protection motor rotation
        .rgxStoppingFault_M[0].2   // Z402.M315B-M1.P51AZ1.Drive feedback error
        .rgxStoppingFault_M[0].15   // Z402.M315B-M2.P51AZ1.Braking resistor anomaly
        .rgxStoppingFault_M[0].4   // Z402.M315B-M1.P403BT1.Motor thermal probe
        .rgxWarning[0].0   // Z402.M315B.Plate not synchronized
        .rgxStoppingFault_M[0].14   // Z402.M315B-M2.P403BT2.Motor thermal probe
        .rgxStoppingFault_M[0].6   // Z402.M315B-M1.Drive not ready
        .rgxStoppingFault_M[0].3   // Z402.M315B-M1.P51AZ1.Local safety switch
        .rgxStoppingFault[0].0   // Z402.M315B.Positioning error
        .rgdFaultCode_M[0]   // Drive fault code M1
        .rgdFaultCode_M[1]   // Drive fault code M2
        .rgxStoppingFault_M[0].5   // Z402.M315B-M1.P51AZ1.Braking resistor anomaly
        .rgxStoppingFault_M[0].16   // Z402.M315B-M2.Drive not ready
        .rgxStoppingFault_M[0].12   // Z402.M315B-M2.P51AZ1.Drive feedback error
        .rgxStoppingFault_M[0].10   // Z402.M315B-M2.P51AZ1.Protection motor rotation
   M315B_Data : UDT_Convoy_SL; {access Read Only}
   M315B_HMR : MAC_Conveyor_HMR := (dState1 := 1, dState3 := 1, dState4 := 1, dStateSensor1 := 1, dStateSensor2 := 1);
        .rgxMan.4   // Run M3 (NU)
        .rgxMan.5   // Reverse M3 (NU)
        .rgxMan.6   // Run M4 (NU)
        .dErrorCode3   // Error code M3 (NU)
        .rgxMan.7   // Reverse M4 (NU)
        .dErrorCode1   // Error code M1
        .rgxMan.0   // Run M1
        .rgxMan.1   // Reverse M1
        .rgxMan.2   // Run M2
        .rgxMan.3   // Reverse M2
        .rgxMan.8   // Run both
        .rgxMan.9   // Reverse both
        .dErrorCode2   // Error code M2
        .dErrorCode4   // Error code M4 (NU)
   M315B_HMW : MAC_Conveyor_HMW;
        .rgxMan.7   // Reverse M4 (NU)
        .rgxMan.5   // Reverse M3 (NU)
        .rgxMan.4   // Run M3 (NU)
        .rgxMan.0   // Run M1
        .rgxMan.1   // Reverse M1
        .rgxMan.2   // Run M2
        .rgxMan.3   // Reverse M2
        .rgxMan.6   // Run M4 (NU)
        .rgxMan.8   // Run both
        .rgxMan.9   // Reverse both
   M315B_M1_DR_IN_MAJ : MOTION_INSTRUCTION := (FLAGS := 570425344, DN := 1); {access None}
   M315B_M1_DR_IN_MAM : MOTION_INSTRUCTION := (FLAGS := 33554432); {access None}
   M315B_M1_DR_IN_MAR : MOTION_INSTRUCTION := (FLAGS := 33554432); {access None}
   M315B_M1_DR_IN_MAS : MOTION_INSTRUCTION := (FLAGS := -1442840576, EN := 1, DN := 1, PC := 1); {access None}
   M315B_M1_DR_IN_MCD : MOTION_INSTRUCTION := (FLAGS := 570425344, DN := 1); {access None}
   M315B_M1_DR_IN_MRP : MOTION_INSTRUCTION := (FLAGS := 33554432); {access None}
   M315B_M1_DR_MAFR : MOTION_INSTRUCTION := (FLAGS := 301989888, ER := 1, ERR := 11); {access None}
   M315B_M1_DR_MDR : MOTION_INSTRUCTION := (FLAGS := -1845493760, EN := 1, ER := 1, ERR := 11); {access None}
   M315B_M1_DR_MSF : MOTION_INSTRUCTION := (FLAGS := 570425344, DN := 1, STATUS := 2, STATE := 1); {access None}
   M315B_M1_DR_MSO : MOTION_INSTRUCTION := (FLAGS := -1610612736, EN := 1, DN := 1, STATE := 1); {access None}
   M315B_M1_DR_OUT_MAJ : MOTION_INSTRUCTION := (FLAGS := 570425344, DN := 1); {access None}
   M315B_M1_DR_OUT_MAM : MOTION_INSTRUCTION := (FLAGS := 33554432); {access None}
   M315B_M1_DR_OUT_MAR : MOTION_INSTRUCTION := (FLAGS := 33554432); {access None}
   M315B_M1_DR_OUT_MAS : MOTION_INSTRUCTION := (FLAGS := -1442840576, EN := 1, DN := 1, PC := 1); {access None}
   M315B_M1_DR_OUT_MCD : MOTION_INSTRUCTION := (FLAGS := 570425344, DN := 1); {access None}
   M315B_M1_DR_OUT_MRP : MOTION_INSTRUCTION := (FLAGS := 33554432); {access None}
   M315B_M2_DR_IN_MAJ : MOTION_INSTRUCTION := (FLAGS := 570425344, DN := 1); {access None}
   M315B_M2_DR_IN_MAM : MOTION_INSTRUCTION := (FLAGS := 33554432); {access None}
   M315B_M2_DR_IN_MAR : MOTION_INSTRUCTION := (FLAGS := 33554432); {access None}
   M315B_M2_DR_IN_MAS : MOTION_INSTRUCTION := (FLAGS := -1442840576, EN := 1, DN := 1, PC := 1); {access None}
   M315B_M2_DR_IN_MCD : MOTION_INSTRUCTION := (FLAGS := 570425344, DN := 1); {access None}
   M315B_M2_DR_IN_MRP : MOTION_INSTRUCTION := (FLAGS := 33554432); {access None}
   M315B_M2_DR_MAFR : MOTION_INSTRUCTION := (FLAGS := 301989888, ER := 1, ERR := 11); {access None}
   M315B_M2_DR_MDR : MOTION_INSTRUCTION := (FLAGS := -1845493760, EN := 1, ER := 1, ERR := 11); {access None}
   M315B_M2_DR_MSF : MOTION_INSTRUCTION := (FLAGS := 570425344, DN := 1, STATUS := 2, STATE := 1); {access None}
   M315B_M2_DR_MSO : MOTION_INSTRUCTION := (FLAGS := -1610612736, EN := 1, DN := 1, STATE := 1); {access None}
   M315B_M2_DR_OUT_MAJ : MOTION_INSTRUCTION := (FLAGS := 570425344, DN := 1); {access None}
   M315B_M2_DR_OUT_MAM : MOTION_INSTRUCTION := (FLAGS := 33554432); {access None}
   M315B_M2_DR_OUT_MAR : MOTION_INSTRUCTION := (FLAGS := 33554432); {access None}
   M315B_M2_DR_OUT_MAS : MOTION_INSTRUCTION := (FLAGS := -1442840576, EN := 1, DN := 1, PC := 1); {access None}
   M315B_M2_DR_OUT_MCD : MOTION_INSTRUCTION := (FLAGS := 570425344, DN := 1); {access None}
   M315B_M2_DR_OUT_MRP : MOTION_INSTRUCTION := (FLAGS := 33554432); {access None}
   M315B_SpaceConv_Utilities : SpaceConv_Utilities := (CONST_dSyncMode := 1, CONST_dSyncroPhWindow_cmm := 450000, CONST_dConveyorLength_cmm := 800000, CONST_dConveyorWidth_cmm := 400000, CONST_dPresetFeedbackTime_ms := 500, CONST_rAcceleration_ms2 := 1.2, CONST_rDeceleration_ms2 := 1.2, CONF_MD1_dScan_ms := 20, CONF_MD2_MD3_dPrstPos_cmm := -390000, CONF_MD4_MD6_dLength_cmm := 365800, CONF_MD7_dOffset_cmm := 50000, ST_dStopLoadForseen_cmm := 620000, ST_dRealSpeed_mm_min := 90000, ST_rStepAdvancementH := 3000.0, ST_rStepAdvancementT := 3000.0, O_xPlateSynchronized := 1, O_dCountFeedbackTime_ms := 500, O_dPresetLoadUnload_cmm := -126300);
   M315B_xOs_PosReq : BOOL;
   M315B_xPlateCullet : BOOL; {access Read Only}
   M315Popup : MAC_Popup_ZC[2] := ([0].ST_xTunnelType := 1, [0].ST_xCleaningConditionOK := 1, [0].ST_xConditionOKForStopCycle := 1, [0].ST_xOutputEnable := 1, [0].ST_xInitialConditionForRise := 1, [0].ST_xExternalConditionToRise := 1, [0].ST_xExternalConditionToDescend := 1, [0].ST_xOutOfEncumbrance := 1, [0].ST_xConditionToReceiveGlass := 1, [0].ST_xEnableControlError := 1, [0].ST_xPlateUnderPopup := 1, [0].ST_xIndexConsPositioning := 1, [0].ST_xPlateComingToPopup := 1, [0].ST_xPlateToBothComing := 1, [0].ST_xPlateToBothPositioning := 1, [0].INPUT_xLiftingProtectionMotor := 1, [0].INPUT_xProtectionCoolingFan := 1, [0].INPUT_xFeedbackCoolingFan := 1, [0].INPUT_xPopupLow := 1, [0].OUTPUT_xPopupVentilation := 1, [0].AUX_dStartPosition_cmm := 4627000, [0].AUX_dEndPosition_cmm := 4827000, [0].AUX_dSpeedConveyor_mm_min := 90000, [0].AUX_dReactionTime_ms := 1500, [0].AUX_dWindowSearch_cmm := 200000, [0].AUX_dDestMaskOpSide := 16#0000_0001, [0].AUX_dReqTarget_cmm := 270000, [0].AUX_dPosPhotocell_cmm := 4627000, [0].AUX_dIndexHead := 3, [0].AUX_dPosTimeout := 5427000, [0].AUX_dIndexPositioning := 3, [0].AUX_dIndexPlateToChangeDestAfterPopup := 1, [0].AUX_tSearchPlateData.dReaction_cmm := 225000, [0].AUX_tSearchPlateData.dPositionDecision_cmm := 4327000, [0].AUX_tSearchPlateData.dPositionStopSearch_cmm := 4627000, [0].AUX_tSearchPlateData.dPositionStopHooked_cmm := 5247000, [0].AUX_tSearchPlateData.dIndex := 3, [0].AUX_tSearchPlateData.xIndexCons := 1, [0].AUX_tSearchPlateData.xPlateHooked := 1, [0].AUX_tSearchPlateData.tResult.rgdHeadPointer[0] := 3, [0].AUX_tSearchPlateData.tResult.rgdHead_cmm[0] := 4328205, [0].AUX_tSearchPlateData.tResult.rgxHead := 1, [0].AUX_tSearchPlateData.tResult.xHeadPresence := 1, [0].tmON_LiftingTimeOut.PRE := 2000, [0].tmON_LiftingFeedbackTimeOut.PRE := 1000, [0].tmOF_WaitBothEndLift.PRE := 1500, [0].tmOF_WaitBothEndLift.ACC := 1500, [0].tmOF_Wait.PRE := 50, [0].tmOF_Wait.ACC := 60, [0].tmON_Saturation.PRE := 1200, [0].tmON_ReentryPlate.PRE := 200, [0].tmON_Positioning.PRE := 40, [1].ST_xTunnelType := 1, [1].ST_xCleaningConditionOK := 1, [1].ST_xConditionOKForStopCycle := 1, [1].ST_xOutputEnable := 1, [1].ST_xInitialConditionForRise := 1, [1].ST_xExternalConditionToRise := 1, [1].ST_xExternalConditionToDescend := 1, [1].ST_xOutOfEncumbrance := 1,
        [1].ST_xConditionToReceiveGlass := 1, [1].ST_xEnableControlError := 1, [1].INPUT_xLiftingProtectionMotor := 1, [1].INPUT_xProtectionCoolingFan := 1, [1].INPUT_xFeedbackCoolingFan := 1, [1].INPUT_xPopupLow := 1, [1].OUTPUT_xPopupVentilation := 1, [1].AUX_dStartPosition_cmm := 4827000, [1].AUX_dEndPosition_cmm := 5027000, [1].AUX_dSpeedConveyor_mm_min := 90000, [1].AUX_dReactionTime_ms := 1500, [1].AUX_dWindowSearch_cmm := 200000, [1].AUX_dDestMaskOpSide := 16#0000_0001, [1].AUX_dPosPhotocell_cmm := 4577000, [1].AUX_dPosTimeout := 5427000, [1].tmON_LiftingTimeOut.PRE := 2000, [1].tmON_LiftingFeedbackTimeOut.PRE := 1000, [1].tmOF_WaitBothEndLift.PRE := 1500, [1].tmOF_WaitBothEndLift.ACC := 1500, [1].tmON_ReentryPlate.PRE := 200, [1].tmON_Positioning.PRE := 40); {access None}
   M315Popup_ALM : MAC_Popup_ZC_ALM[2]; {access Read Only}
        [0].rgxFault[0].0   // M315PopupUP.Lifting protection motor
        [0].rgxFault[0].1   // M315PopupUP.Lifting feedback motor
        [0].rgxFault[0].3   // M315PopupUP.Lifting fan protection
        [0].rgxFault[0].4   // M315PopupUP.Lifting fan feedback
        [0].rgxFault[0].2   // M315PopupUP.Lifting safety switch
        [1].rgxFault[0].0   // M315PopupDN.Lifting protection motor
        [1].rgxFault[0].1   // M315PopupDN.Lifting feedback motor
        [1].rgxFault[0].3   // M315PopupDN.Lifting fan protection
        [1].rgxFault[0].4   // M315PopupDN.Lifting fan feedback
        [1].rgxWarning[0].0   // M315PopupDN.Positioning error on conveyor
        [1].rgxFault[0].2   // M315PopupDN.Lifting safety switch
        [1].rgxStoppingFault[0].0   // M315PopupDN.Lifting position error
        [0].rgxWarning[0].0   // M315PopupUP.Positioning error on conveyor
        [0].rgxStoppingFault[0].0   // M315PopupUP.Lifting position error
   M315Popup_HMR : MAC_Popup_ZC_HMR[2] := ([0].xHighPosition := 1, [0].rgdState := 1, [1].xHighPosition := 1, [1].rgdState := 1); {access Read Only}
        [0].rgxMan.0   // Rise popup upstream {x|x|x|x|O}
        [0].rgxMan.1   // Lower popup upstream {x|x|x|x|O}
        [0].rgxMan.2   // Rise both popup {x|x|x|x|O}
        [0].rgxMan.3   // Lower both popup {x|x|x|x|O}
        [1].rgxMan.0   // Rise popup downstream {x|x|x|x|O}
        [1].rgxMan.1   // Lower popup downstream {x|x|x|x|O}
   M315Popup_HMW : MAC_Popup_ZC_HMW[2] := ([0].dSingleCapOffset_cmm := 20000, [0].dSaturationSelection := 2);
        [0].rgxMan.0   // Rise popup upstream {x|x|x|x|O}
        [0].rgxMan.1   // Lower popup upstream {x|x|x|x|O}
        [0].rgxMan.2   // Rise both popup {x|x|x|x|O}
        [0].rgxMan.3   // Lower both popup {x|x|x|x|O}
        [1].rgxMan.0   // Rise popup downstream {x|x|x|x|O}
        [1].rgxMan.1   // Lower popup downstream {x|x|x|x|O}
   M315Popup_IN_MOTION : MAC_Popup_ZC_IN_MOTION[2]; {access None}
   M315Popup_OUT_MOTION : MAC_Popup_ZC_OUT_MOTION[2]; {access None}
   M315Popup_PlateFreeTimeout : TIMER; {access Read Only}
   M315Popup_ReentryCap : UDT_ConvoyCap_ZC;
   M315Popup_SL_DATA : UDT_Convoy_SL;
   M315Popup_tSearchPlateChangeFromCS4402 : GP_TrackingSearchPlate_STC; {access Read Only}
   M315Popup_xDrivePosEnable : BOOL; {access Read Only}
   M315Popup_xEndRise : BOOL; {access Read Only}
   M315Popup_xEndRiseWaitingForCondition : BOOL; {access Read Only}
   M316 : MAC_Conveyor := (ST_xCleaningConditionOK := 1, ST_xEnableControlError := 1, ST_xPlateSynchronized := 1, ST_xSafetyMovement := 1, OSR_xSynchroPhotocellTail := 1, INPUT_xDriveReady_M1 := 1, INPUT_xLocalSafetySwitch_M1 := 1, INPUT_xMotorThermalProbe_M1 := 1, INPUT_xProtectionMotor_M1 := 1, INPUT_xDriveReady_M2 := 1, INPUT_xLocalSafetySwitch_M2 := 1, INPUT_xMotorThermalProbe_M2 := 1, INPUT_xProtectionMotor_M2 := 1, OUTPUT_xDriveEnable_M1 := 1, OUTPUT_xDriveEnable_M2 := 1, AUX_dPresetStopLoad_cmm := 408333, AUX_dPresetStopUnload_cmm := 491667, AUX_dAccSpace_cmm := 41667, AUX_dDecSpace_cmm := 41667, AUX_dReqSpeed_mm_min := 60000, AUX_dPhPosTarget_cmm := 295000, AUX_dPhPosTarget_2_cmm := 169750, tmON_FeedbackTimeOut_M1.PRE := 1500, tmOF_DriveEnable_M1.PRE := 30000, tmOF_DriveEnable_M1.ACC := 1820, tmOF_DriveEnable_M1.TT := 1, tmOF_DriveEnable_M1.DN := 1, tmOF_PowerSaving_M1.PRE := 20000, tmOF_PowerSaving_M1.ACC := 20000, tmON_FeedbackTimeOut_M2.PRE := 2000, tmOF_DriveEnable_M2.PRE := 30000, tmOF_DriveEnable_M2.ACC := 1820, tmOF_DriveEnable_M2.TT := 1, tmOF_DriveEnable_M2.DN := 1, tmOF_PowerSaving_M2.PRE := 20000, tmON_AuxFunction6.PRE := 5000, tmON_AuxFunction7.PRE := 100, tmON_AuxFunction8.PRE := 100, tmOF_MCD_M1.PRE := 200, tmOF_MCD_M1.ACC := 200, tmOF_MCD_M2.PRE := 200, tmOF_MCD_M2.ACC := 200); {access None}
        .INPUT_xMotorThermalProbe_M2   // M403.M2.P403BT4. Motor thermal probe
        .ST_xAux1   // request rise popup to unload on M325 (reentry)
        .INPUT_xMotorThermalProbe_M1   // M403.M1.P403BT3. Motor thermal probe